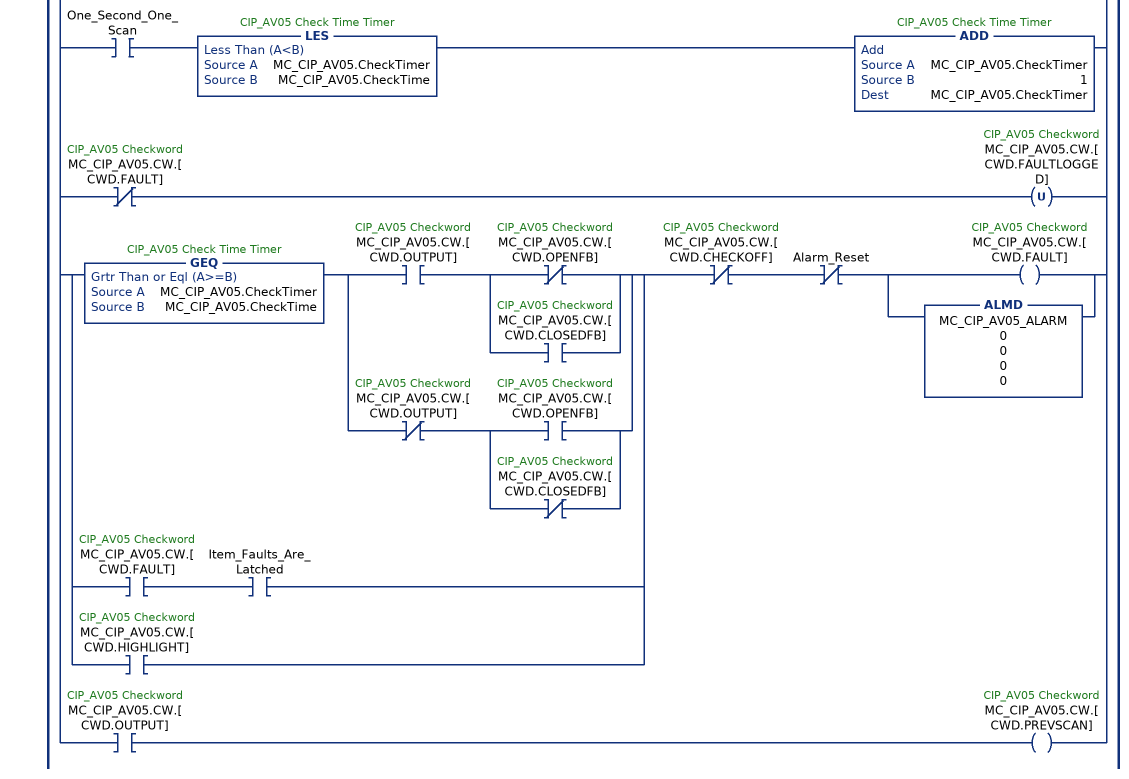
   62: [NEQ(MC_CIP_AV05.DriveBits,0) OTE(MC_CIP_AV05.CW.[CWD.AUTODRV]) ,[XIC(MC_CIP_AV05.CW.[CWD.AUTODRV]) XIO(MC_CIP_AV05.CW.[CWD.MANUAL]) ,XIC(MC_CIP_AV05.CW.[CWD.MANDRV]) XIC(MC_CIP_AV05.CW.[CWD.MANUAL]) ] OTE(MC_CIP_AV05.CW.[CWD.OUTPUT]) ,XIC(MC_CIP_AV05.CW.[CWD.OUTPUT]) OTE(MC_CIP_AV05_DR) ,XIC(S:FS) [OTU(MC_CIP_AV05.CW.[CWD.MANUAL]) ,LEQ(MC_CIP_AV05.CheckTime,0) MOV(Default_Check_Time,MC_CIP_AV05.CheckTime) ] ,[[XIC(MC_CIP_AV05_O) XIO(Item_Simulation_Flag) ,XIC(Item_Simulation_Flag) XIC(MC_CIP_AV05.CW.[CWD.OUTPUT]) XIO(MC_CIP_AV05.CW.[CWD.SIMFAIL]) ] OTE(MC_CIP_AV05.CW.[CWD.OPENFB]) ,[XIC(MC_CIP_AV05_C) XIO(Item_Simulation_Flag) ,XIC(Item_Simulation_Flag) XIO(MC_CIP_AV05.CW.[CWD.OUTPUT]) XIO(MC_CIP_AV05.CW.[CWD.SIMFAIL]) ] OTE(MC_CIP_AV05.CW.[CWD.CLOSEDFB]) ] ,[XIC(MC_CIP_AV05.CW.[CWD.OUTPUT]) XIO(MC_CIP_AV05.CW.[CWD.PREVSCAN]) ,XIO(MC_CIP_AV05.CW.[CWD.OUTPUT]) XIC(MC_CIP_AV05.CW.[CWD.PREVSCAN]) ] CLR(MC_CIP_AV05.CheckTimer) ,XIC(One_Second_One_Scan) LES(MC_CIP_AV05.CheckTimer,MC_CIP_AV05.CheckTime) ADD(MC_CIP_AV05.CheckTimer,1,MC_CIP_AV05.CheckTimer) ,XIO(MC_CIP_AV05.CW.[CWD.FAULT]) OTU(MC_CIP_AV05.CW.[CWD.FAULTLOGGED]) ,[GEQ(MC_CIP_AV05.CheckTimer,MC_CIP_AV05.CheckTime) [XIC(MC_CIP_AV05.CW.[CWD.OUTPUT]) [XIO(MC_CIP_AV05.CW.[CWD.OPENFB]) ,XIC(MC_CIP_AV05.CW.[CWD.CLOSEDFB]) ] ,XIO(MC_CIP_AV05.CW.[CWD.OUTPUT]) [XIC(MC_CIP_AV05.CW.[CWD.OPENFB]) ,XIO(MC_CIP_AV05.CW.[CWD.CLOSEDFB]) ] ] ,XIC(MC_CIP_AV05.CW.[CWD.FAULT]) XIC(Item_Faults_Are_Latched) ,XIC(MC_CIP_AV05.CW.[CWD.HIGHLIGHT]) ] XIO(MC_CIP_AV05.CW.[CWD.CHECKOFF]) XIO(Alarm_Reset) [OTE(MC_CIP_AV05.CW.[CWD.FAULT]) ,ALMD(MC_CIP_AV05_ALARM,0,0,0,0) ] ,XIC(MC_CIP_AV05.CW.[CWD.OUTPUT]) OTE(MC_CIP_AV05.CW.[CWD.PREVSCAN]) ];
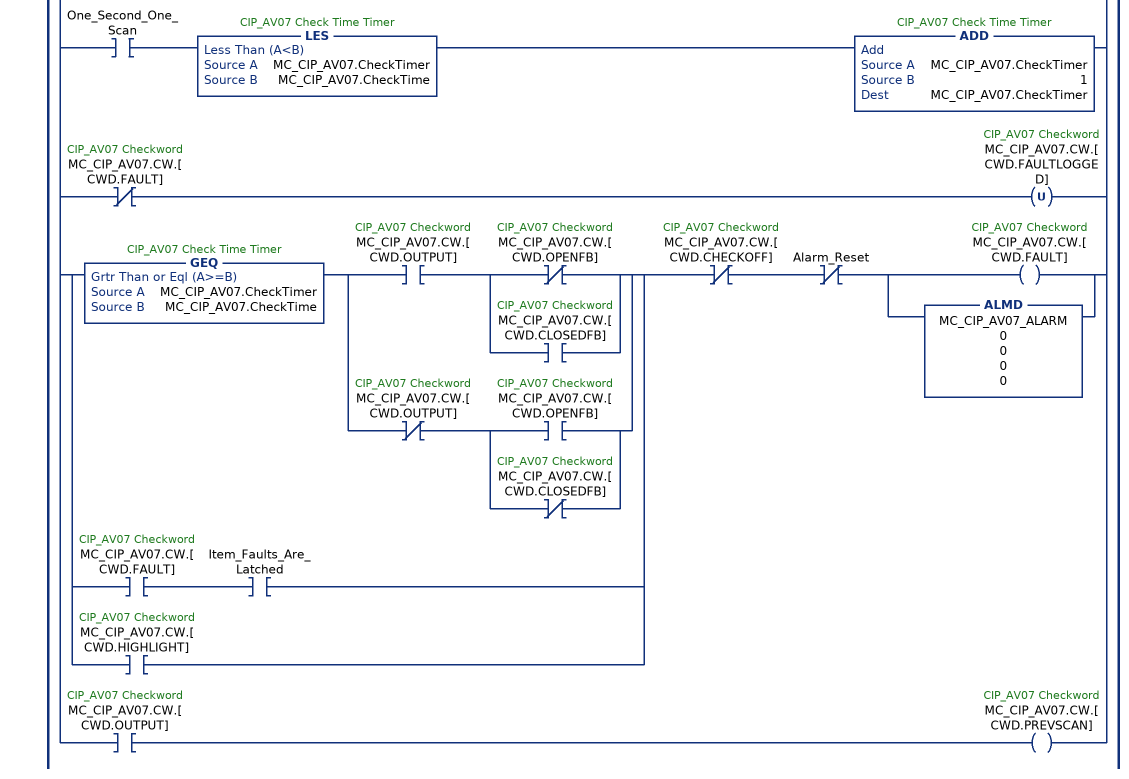
   63: [NEQ(MC_CIP_AV07.DriveBits,0) OTE(MC_CIP_AV07.CW.[CWD.AUTODRV]) ,[XIC(MC_CIP_AV07.CW.[CWD.AUTODRV]) XIO(MC_CIP_AV07.CW.[CWD.MANUAL]) ,XIC(MC_CIP_AV07.CW.[CWD.MANDRV]) XIC(MC_CIP_AV07.CW.[CWD.MANUAL]) ] OTE(MC_CIP_AV07.CW.[CWD.OUTPUT]) ,XIC(MC_CIP_AV07.CW.[CWD.OUTPUT]) OTE(MC_CIP_AV07_DR) ,XIC(S:FS) [OTU(MC_CIP_AV07.CW.[CWD.MANUAL]) ,LEQ(MC_CIP_AV07.CheckTime,0) MOV(Default_Check_Time,MC_CIP_AV07.CheckTime) ] ,[[XIC(MC_CIP_AV07_O) XIO(Item_Simulation_Flag) ,XIC(Item_Simulation_Flag) XIC(MC_CIP_AV07.CW.[CWD.OUTPUT]) XIO(MC_CIP_AV07.CW.[CWD.SIMFAIL]) ] OTE(MC_CIP_AV07.CW.[CWD.OPENFB]) ,[XIC(MC_CIP_AV07_C) XIO(Item_Simulation_Flag) ,XIC(Item_Simulation_Flag) XIO(MC_CIP_AV07.CW.[CWD.OUTPUT]) XIO(MC_CIP_AV07.CW.[CWD.SIMFAIL]) ] OTE(MC_CIP_AV07.CW.[CWD.CLOSEDFB]) ] ,[XIC(MC_CIP_AV07.CW.[CWD.OUTPUT]) XIO(MC_CIP_AV07.CW.[CWD.PREVSCAN]) ,XIO(MC_CIP_AV07.CW.[CWD.OUTPUT]) XIC(MC_CIP_AV07.CW.[CWD.PREVSCAN]) ] CLR(MC_CIP_AV07.CheckTimer) ,XIC(One_Second_One_Scan) LES(MC_CIP_AV07.CheckTimer,MC_CIP_AV07.CheckTime) ADD(MC_CIP_AV07.CheckTimer,1,MC_CIP_AV07.CheckTimer) ,XIO(MC_CIP_AV07.CW.[CWD.FAULT]) OTU(MC_CIP_AV07.CW.[CWD.FAULTLOGGED]) ,[GEQ(MC_CIP_AV07.CheckTimer,MC_CIP_AV07.CheckTime) [XIC(MC_CIP_AV07.CW.[CWD.OUTPUT]) [XIO(MC_CIP_AV07.CW.[CWD.OPENFB]) ,XIC(MC_CIP_AV07.CW.[CWD.CLOSEDFB]) ] ,XIO(MC_CIP_AV07.CW.[CWD.OUTPUT]) [XIC(MC_CIP_AV07.CW.[CWD.OPENFB]) ,XIO(MC_CIP_AV07.CW.[CWD.CLOSEDFB]) ] ] ,XIC(MC_CIP_AV07.CW.[CWD.FAULT]) XIC(Item_Faults_Are_Latched) ,XIC(MC_CIP_AV07.CW.[CWD.HIGHLIGHT]) ] XIO(MC_CIP_AV07.CW.[CWD.CHECKOFF]) XIO(Alarm_Reset) [OTE(MC_CIP_AV07.CW.[CWD.FAULT]) ,ALMD(MC_CIP_AV07_ALARM,0,0,0,0) ] ,XIC(MC_CIP_AV07.CW.[CWD.OUTPUT]) OTE(MC_CIP_AV07.CW.[CWD.PREVSCAN]) ];
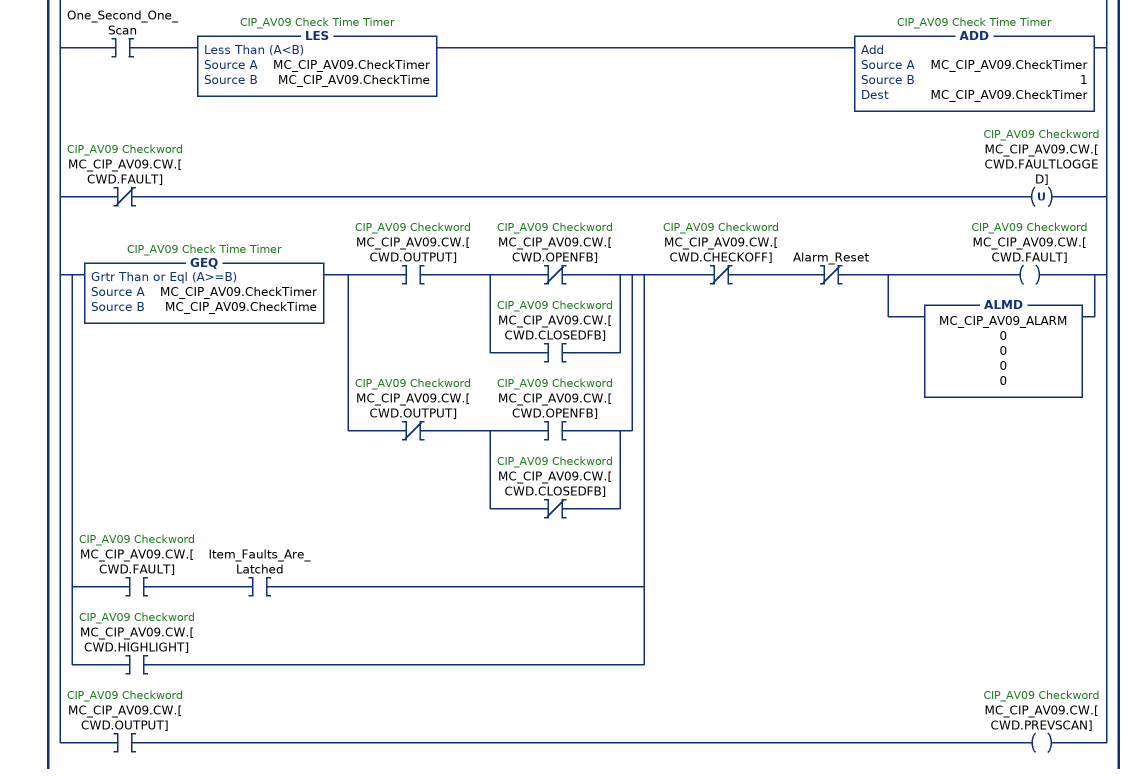
   64: [NEQ(MC_CIP_AV09.DriveBits,0) OTE(MC_CIP_AV09.CW.[CWD.AUTODRV]) ,[XIC(MC_CIP_AV09.CW.[CWD.AUTODRV]) XIO(MC_CIP_AV09.CW.[CWD.MANUAL]) ,XIC(MC_CIP_AV09.CW.[CWD.MANDRV]) XIC(MC_CIP_AV09.CW.[CWD.MANUAL]) ] OTE(MC_CIP_AV09.CW.[CWD.OUTPUT]) ,XIC(MC_CIP_AV09.CW.[CWD.OUTPUT]) OTE(MC_CIP_AV09_DR) ,XIC(S:FS) [OTU(MC_CIP_AV09.CW.[CWD.MANUAL]) ,LEQ(MC_CIP_AV09.CheckTime,0) MOV(Default_Check_Time,MC_CIP_AV09.CheckTime) ] ,[[XIC(MC_CIP_AV09_O) XIO(Item_Simulation_Flag) ,XIC(Item_Simulation_Flag) XIC(MC_CIP_AV09.CW.[CWD.OUTPUT]) XIO(MC_CIP_AV09.CW.[CWD.SIMFAIL]) ] OTE(MC_CIP_AV09.CW.[CWD.OPENFB]) ,[XIC(MC_CIP_AV09_C) XIO(Item_Simulation_Flag) ,XIC(Item_Simulation_Flag) XIO(MC_CIP_AV09.CW.[CWD.OUTPUT]) XIO(MC_CIP_AV09.CW.[CWD.SIMFAIL]) ] OTE(MC_CIP_AV09.CW.[CWD.CLOSEDFB]) ] ,[XIC(MC_CIP_AV09.CW.[CWD.OUTPUT]) XIO(MC_CIP_AV09.CW.[CWD.PREVSCAN]) ,XIO(MC_CIP_AV09.CW.[CWD.OUTPUT]) XIC(MC_CIP_AV09.CW.[CWD.PREVSCAN]) ] CLR(MC_CIP_AV09.CheckTimer) ,XIC(One_Second_One_Scan) LES(MC_CIP_AV09.CheckTimer,MC_CIP_AV09.CheckTime) ADD(MC_CIP_AV09.CheckTimer,1,MC_CIP_AV09.CheckTimer) ,XIO(MC_CIP_AV09.CW.[CWD.FAULT]) OTU(MC_CIP_AV09.CW.[CWD.FAULTLOGGED]) ,[GEQ(MC_CIP_AV09.CheckTimer,MC_CIP_AV09.CheckTime) [XIC(MC_CIP_AV09.CW.[CWD.OUTPUT]) [XIO(MC_CIP_AV09.CW.[CWD.OPENFB]) ,XIC(MC_CIP_AV09.CW.[CWD.CLOSEDFB]) ] ,XIO(MC_CIP_AV09.CW.[CWD.OUTPUT]) [XIC(MC_CIP_AV09.CW.[CWD.OPENFB]) ,XIO(MC_CIP_AV09.CW.[CWD.CLOSEDFB]) ] ] ,XIC(MC_CIP_AV09.CW.[CWD.FAULT]) XIC(Item_Faults_Are_Latched) ,XIC(MC_CIP_AV09.CW.[CWD.HIGHLIGHT]) ] XIO(MC_CIP_AV09.CW.[CWD.CHECKOFF]) XIO(Alarm_Reset) [OTE(MC_CIP_AV09.CW.[CWD.FAULT]) ,ALMD(MC_CIP_AV09_ALARM,0,0,0,0) ] ,XIC(MC_CIP_AV09.CW.[CWD.OUTPUT]) OTE(MC_CIP_AV09.CW.[CWD.PREVSCAN]) ];
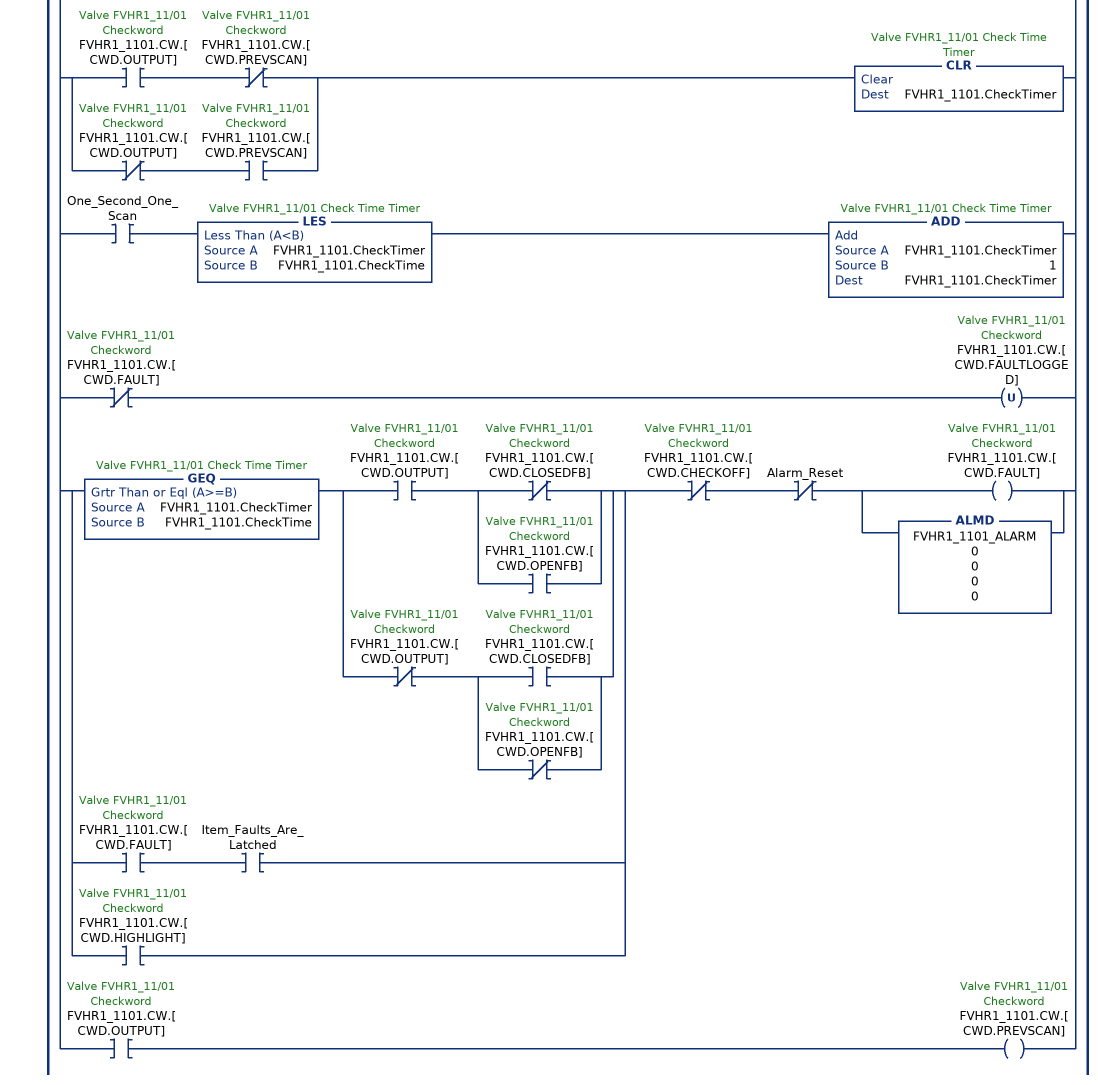
   65: [NEQ(FVHR1_1101.DriveBits,0) OTE(FVHR1_1101.CW.[CWD.AUTODRV]) ,[XIC(FVHR1_1101.CW.[CWD.AUTODRV]) XIO(FVHR1_1101.CW.[CWD.MANUAL]) ,XIC(FVHR1_1101.CW.[CWD.MANDRV]) XIC(FVHR1_1101.CW.[CWD.MANUAL]) ] OTE(FVHR1_1101.CW.[CWD.OUTPUT]) ,XIC(FVHR1_1101.CW.[CWD.OUTPUT]) OTE(FVHR1_1101_DR) ,XIC(S:FS) [OTU(FVHR1_1101.CW.[CWD.MANUAL]) ,LEQ(FVHR1_1101.CheckTime,0) MOV(Default_Check_Time,FVHR1_1101.CheckTime) ] ,[[XIC(FVHR1_1101_OP) XIO(Item_Simulation_Flag) ,XIC(Item_Simulation_Flag) XIC(FVHR1_1101.CW.[CWD.OUTPUT]) XIO(FVHR1_1101.CW.[CWD.SIMFAIL]) ] OTE(FVHR1_1101.CW.[CWD.OPENFB]) ,[XIC(FVHR1_1101_CL) XIO(Item_Simulation_Flag) ,XIC(Item_Simulation_Flag) XIO(FVHR1_1101.CW.[CWD.OUTPUT]) XIO(FVHR1_1101.CW.[CWD.SIMFAIL]) ] OTE(FVHR1_1101.CW.[CWD.CLOSEDFB]) ] ,[XIC(FVHR1_1101.CW.[CWD.OUTPUT]) XIO(FVHR1_1101.CW.[CWD.PREVSCAN]) ,XIO(FVHR1_1101.CW.[CWD.OUTPUT]) XIC(FVHR1_1101.CW.[CWD.PREVSCAN]) ] CLR(FVHR1_1101.CheckTimer) ,XIC(One_Second_One_Scan) LES(FVHR1_1101.CheckTimer,FVHR1_1101.CheckTime) ADD(FVHR1_1101.CheckTimer,1,FVHR1_1101.CheckTimer) ,XIO(FVHR1_1101.CW.[CWD.FAULT]) OTU(FVHR1_1101.CW.[CWD.FAULTLOGGED]) ,[GEQ(FVHR1_1101.CheckTimer,FVHR1_1101.CheckTime) [XIC(FVHR1_1101.CW.[CWD.OUTPUT]) [XIO(FVHR1_1101.CW.[CWD.CLOSEDFB]) ,XIC(FVHR1_1101.CW.[CWD.OPENFB]) ] ,XIO(FVHR1_1101.CW.[CWD.OUTPUT]) [XIC(FVHR1_1101.CW.[CWD.CLOSEDFB]) ,XIO(FVHR1_1101.CW.[CWD.OPENFB]) ] ] ,XIC(FVHR1_1101.CW.[CWD.FAULT]) XIC(Item_Faults_Are_Latched) ,XIC(FVHR1_1101.CW.[CWD.HIGHLIGHT]) ] XIO(FVHR1_1101.CW.[CWD.CHECKOFF]) XIO(Alarm_Reset) [OTE(FVHR1_1101.CW.[CWD.FAULT]) ,ALMD(FVHR1_1101_ALARM,0,0,0,0) ] ,XIC(FVHR1_1101.CW.[CWD.OUTPUT]) OTE(FVHR1_1101.CW.[CWD.PREVSCAN]) ];
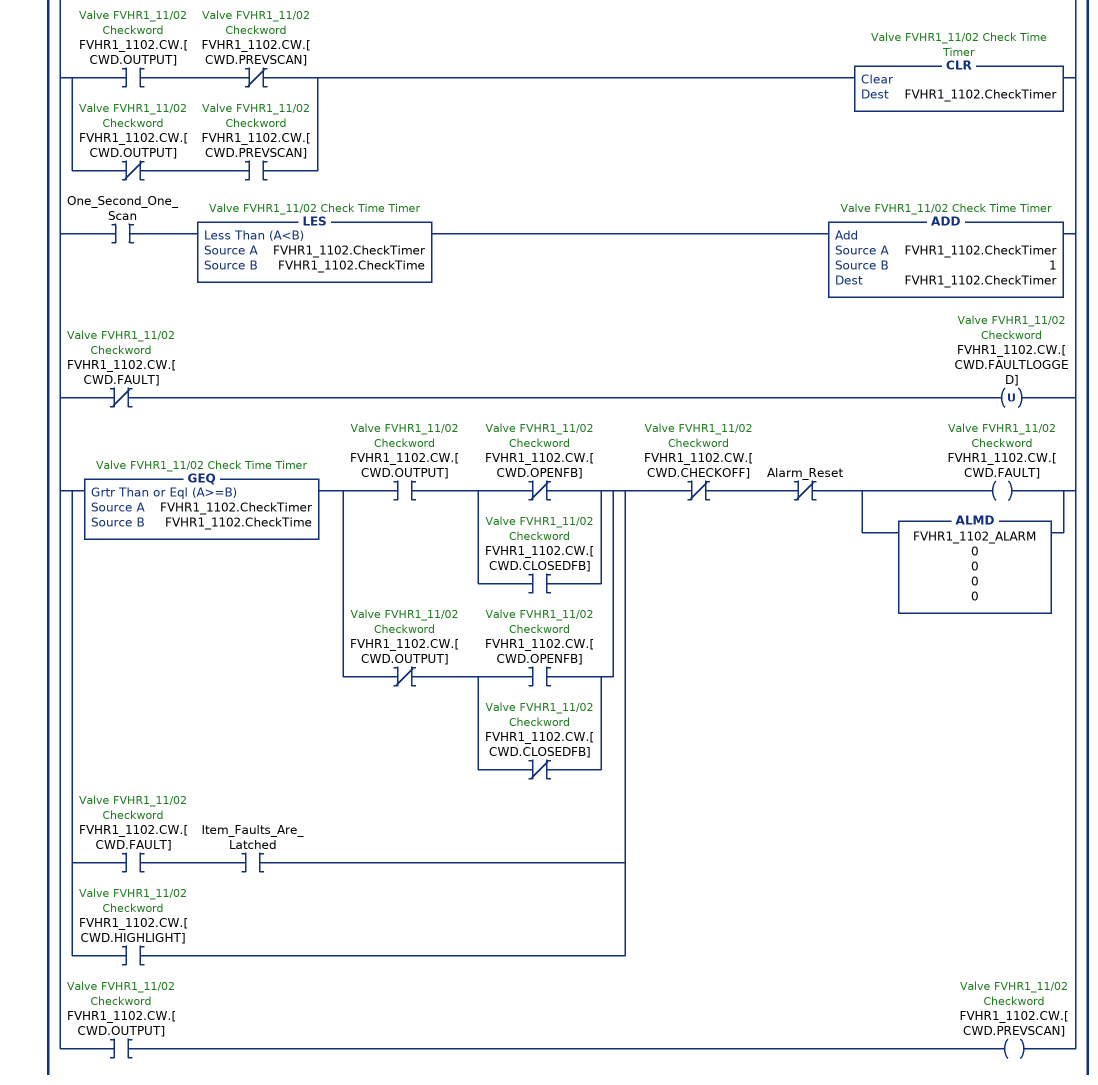
   66: [NEQ(FVHR1_1102.DriveBits,0) OTE(FVHR1_1102.CW.[CWD.AUTODRV]) ,[XIC(FVHR1_1102.CW.[CWD.AUTODRV]) XIO(FVHR1_1102.CW.[CWD.MANUAL]) ,XIC(FVHR1_1102.CW.[CWD.MANDRV]) XIC(FVHR1_1102.CW.[CWD.MANUAL]) ] OTE(FVHR1_1102.CW.[CWD.OUTPUT]) ,XIC(FVHR1_1102.CW.[CWD.OUTPUT]) OTE(FVHR1_1102_DR) ,XIC(S:FS) [OTU(FVHR1_1102.CW.[CWD.MANUAL]) ,LEQ(FVHR1_1102.CheckTime,0) MOV(Default_Check_Time,FVHR1_1102.CheckTime) ] ,[[XIC(FVHR1_1102_OP) XIO(Item_Simulation_Flag) ,XIC(Item_Simulation_Flag) XIC(FVHR1_1102.CW.[CWD.OUTPUT]) XIO(FVHR1_1102.CW.[CWD.SIMFAIL]) ] OTE(FVHR1_1102.CW.[CWD.OPENFB]) ,[XIC(FVHR1_1102_CL) XIO(Item_Simulation_Flag) ,XIC(Item_Simulation_Flag) XIO(FVHR1_1102.CW.[CWD.OUTPUT]) XIO(FVHR1_1102.CW.[CWD.SIMFAIL]) ] OTE(FVHR1_1102.CW.[CWD.CLOSEDFB]) ] ,[XIC(FVHR1_1102.CW.[CWD.OUTPUT]) XIO(FVHR1_1102.CW.[CWD.PREVSCAN]) ,XIO(FVHR1_1102.CW.[CWD.OUTPUT]) XIC(FVHR1_1102.CW.[CWD.PREVSCAN]) ] CLR(FVHR1_1102.CheckTimer) ,XIC(One_Second_One_Scan) LES(FVHR1_1102.CheckTimer,FVHR1_1102.CheckTime) ADD(FVHR1_1102.CheckTimer,1,FVHR1_1102.CheckTimer) ,XIO(FVHR1_1102.CW.[CWD.FAULT]) OTU(FVHR1_1102.CW.[CWD.FAULTLOGGED]) ,[GEQ(FVHR1_1102.CheckTimer,FVHR1_1102.CheckTime) [XIC(FVHR1_1102.CW.[CWD.OUTPUT]) [XIO(FVHR1_1102.CW.[CWD.OPENFB]) ,XIC(FVHR1_1102.CW.[CWD.CLOSEDFB]) ] ,XIO(FVHR1_1102.CW.[CWD.OUTPUT]) [XIC(FVHR1_1102.CW.[CWD.OPENFB]) ,XIO(FVHR1_1102.CW.[CWD.CLOSEDFB]) ] ] ,XIC(FVHR1_1102.CW.[CWD.FAULT]) XIC(Item_Faults_Are_Latched) ,XIC(FVHR1_1102.CW.[CWD.HIGHLIGHT]) ] XIO(FVHR1_1102.CW.[CWD.CHECKOFF]) XIO(Alarm_Reset) [OTE(FVHR1_1102.CW.[CWD.FAULT]) ,ALMD(FVHR1_1102_ALARM,0,0,0,0) ] ,XIC(FVHR1_1102.CW.[CWD.OUTPUT]) OTE(FVHR1_1102.CW.[CWD.PREVSCAN]) ];
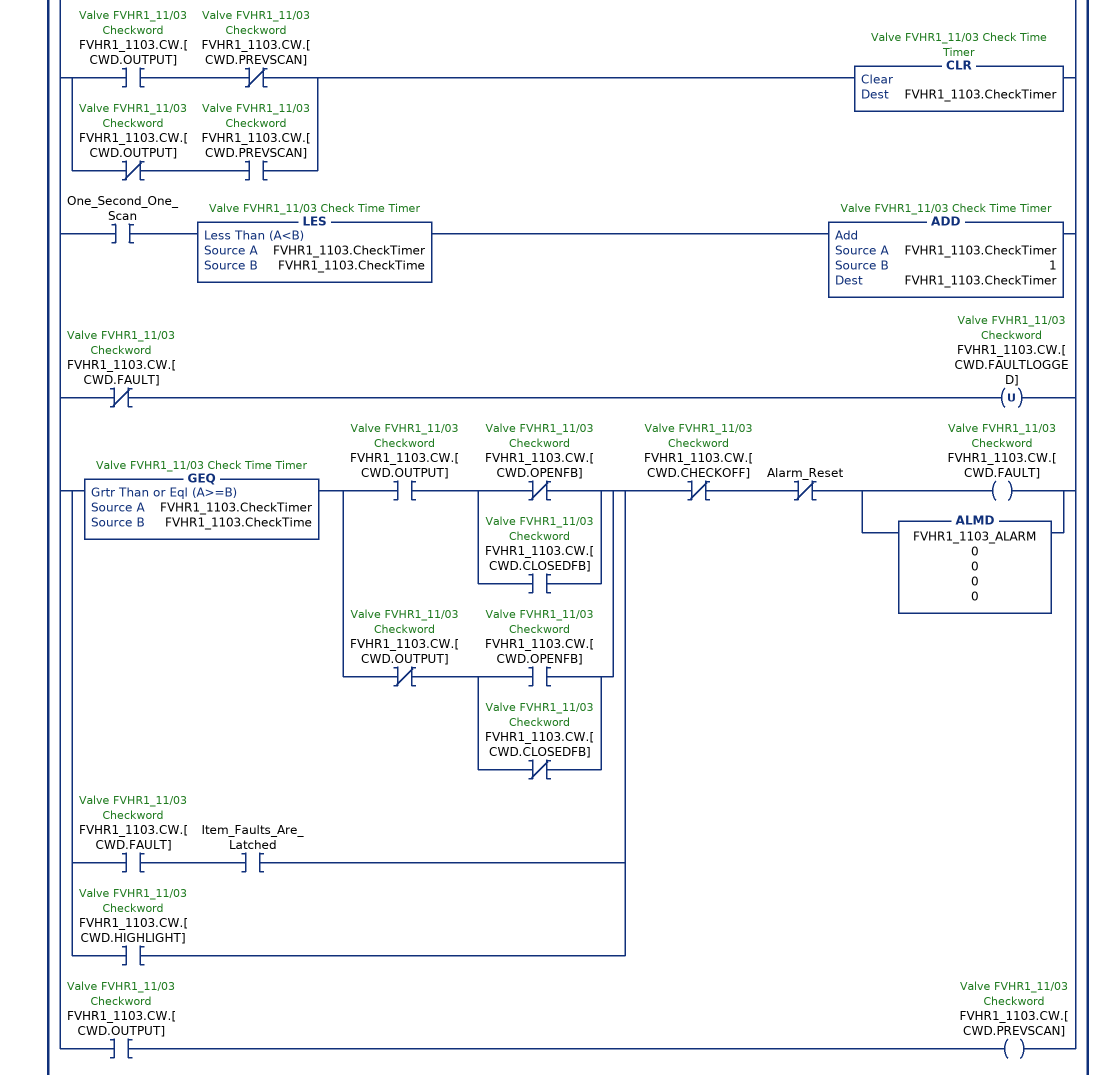
   67: [NEQ(FVHR1_1103.DriveBits,0) OTE(FVHR1_1103.CW.[CWD.AUTODRV]) ,[XIC(FVHR1_1103.CW.[CWD.AUTODRV]) XIO(FVHR1_1103.CW.[CWD.MANUAL]) ,XIC(FVHR1_1103.CW.[CWD.MANDRV]) XIC(FVHR1_1103.CW.[CWD.MANUAL]) ] OTE(FVHR1_1103.CW.[CWD.OUTPUT]) ,XIC(FVHR1_1103.CW.[CWD.OUTPUT]) OTE(FVHR1_1103_DR) ,XIC(S:FS) [OTU(FVHR1_1103.CW.[CWD.MANUAL]) ,LEQ(FVHR1_1103.CheckTime,0) MOV(Default_Check_Time,FVHR1_1103.CheckTime) ] ,[[XIC(FVHR1_1103_OP) XIO(Item_Simulation_Flag) ,XIC(Item_Simulation_Flag) XIC(FVHR1_1103.CW.[CWD.OUTPUT]) XIO(FVHR1_1103.CW.[CWD.SIMFAIL]) ] OTE(FVHR1_1103.CW.[CWD.OPENFB]) ,[XIC(FVHR1_1103_CL) XIO(Item_Simulation_Flag) ,XIC(Item_Simulation_Flag) XIO(FVHR1_1103.CW.[CWD.OUTPUT]) XIO(FVHR1_1103.CW.[CWD.SIMFAIL]) ] OTE(FVHR1_1103.CW.[CWD.CLOSEDFB]) ] ,[XIC(FVHR1_1103.CW.[CWD.OUTPUT]) XIO(FVHR1_1103.CW.[CWD.PREVSCAN]) ,XIO(FVHR1_1103.CW.[CWD.OUTPUT]) XIC(FVHR1_1103.CW.[CWD.PREVSCAN]) ] CLR(FVHR1_1103.CheckTimer) ,XIC(One_Second_One_Scan) LES(FVHR1_1103.CheckTimer,FVHR1_1103.CheckTime) ADD(FVHR1_1103.CheckTimer,1,FVHR1_1103.CheckTimer) ,XIO(FVHR1_1103.CW.[CWD.FAULT]) OTU(FVHR1_1103.CW.[CWD.FAULTLOGGED]) ,[GEQ(FVHR1_1103.CheckTimer,FVHR1_1103.CheckTime) [XIC(FVHR1_1103.CW.[CWD.OUTPUT]) [XIO(FVHR1_1103.CW.[CWD.OPENFB]) ,XIC(FVHR1_1103.CW.[CWD.CLOSEDFB]) ] ,XIO(FVHR1_1103.CW.[CWD.OUTPUT]) [XIC(FVHR1_1103.CW.[CWD.OPENFB]) ,XIO(FVHR1_1103.CW.[CWD.CLOSEDFB]) ] ] ,XIC(FVHR1_1103.CW.[CWD.FAULT]) XIC(Item_Faults_Are_Latched) ,XIC(FVHR1_1103.CW.[CWD.HIGHLIGHT]) ] XIO(FVHR1_1103.CW.[CWD.CHECKOFF]) XIO(Alarm_Reset) [OTE(FVHR1_1103.CW.[CWD.FAULT]) ,ALMD(FVHR1_1103_ALARM,0,0,0,0) ] ,XIC(FVHR1_1103.CW.[CWD.OUTPUT]) OTE(FVHR1_1103.CW.[CWD.PREVSCAN]) ];
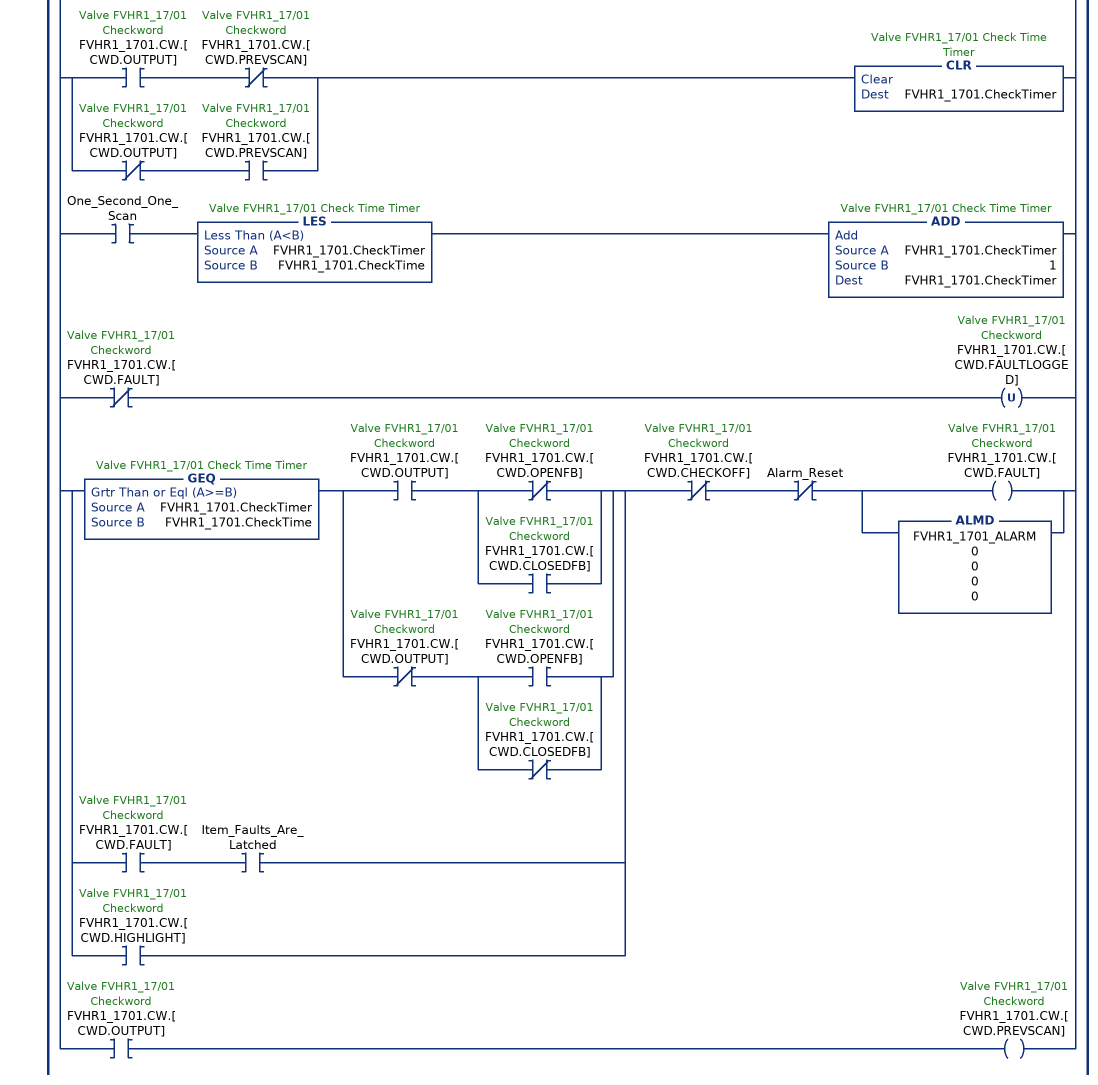
   68: [NEQ(FVHR1_1701.DriveBits,0) OTE(FVHR1_1701.CW.[CWD.AUTODRV]) ,[XIC(FVHR1_1701.CW.[CWD.AUTODRV]) XIO(FVHR1_1701.CW.[CWD.MANUAL]) ,XIC(FVHR1_1701.CW.[CWD.MANDRV]) XIC(FVHR1_1701.CW.[CWD.MANUAL]) ] OTE(FVHR1_1701.CW.[CWD.OUTPUT]) ,XIC(FVHR1_1701.CW.[CWD.OUTPUT]) OTE(FVHR1_1701_DR) ,XIC(S:FS) [OTU(FVHR1_1701.CW.[CWD.MANUAL]) ,LEQ(FVHR1_1701.CheckTime,0) MOV(Default_Check_Time,FVHR1_1701.CheckTime) ] ,[[XIC(FVHR1_1701_OP) XIO(Item_Simulation_Flag) ,XIC(Item_Simulation_Flag) XIC(FVHR1_1701.CW.[CWD.OUTPUT]) XIO(FVHR1_1701.CW.[CWD.SIMFAIL]) ] OTE(FVHR1_1701.CW.[CWD.OPENFB]) ,[XIC(FVHR1_1701_CL) XIO(Item_Simulation_Flag) ,XIC(Item_Simulation_Flag) XIO(FVHR1_1701.CW.[CWD.OUTPUT]) XIO(FVHR1_1701.CW.[CWD.SIMFAIL]) ] OTE(FVHR1_1701.CW.[CWD.CLOSEDFB]) ] ,[XIC(FVHR1_1701.CW.[CWD.OUTPUT]) XIO(FVHR1_1701.CW.[CWD.PREVSCAN]) ,XIO(FVHR1_1701.CW.[CWD.OUTPUT]) XIC(FVHR1_1701.CW.[CWD.PREVSCAN]) ] CLR(FVHR1_1701.CheckTimer) ,XIC(One_Second_One_Scan) LES(FVHR1_1701.CheckTimer,FVHR1_1701.CheckTime) ADD(FVHR1_1701.CheckTimer,1,FVHR1_1701.CheckTimer) ,XIO(FVHR1_1701.CW.[CWD.FAULT]) OTU(FVHR1_1701.CW.[CWD.FAULTLOGGED]) ,[GEQ(FVHR1_1701.CheckTimer,FVHR1_1701.CheckTime) [XIC(FVHR1_1701.CW.[CWD.OUTPUT]) [XIO(FVHR1_1701.CW.[CWD.OPENFB]) ,XIC(FVHR1_1701.CW.[CWD.CLOSEDFB]) ] ,XIO(FVHR1_1701.CW.[CWD.OUTPUT]) [XIC(FVHR1_1701.CW.[CWD.OPENFB]) ,XIO(FVHR1_1701.CW.[CWD.CLOSEDFB]) ] ] ,XIC(FVHR1_1701.CW.[CWD.FAULT]) XIC(Item_Faults_Are_Latched) ,XIC(FVHR1_1701.CW.[CWD.HIGHLIGHT]) ] XIO(FVHR1_1701.CW.[CWD.CHECKOFF]) XIO(Alarm_Reset) [OTE(FVHR1_1701.CW.[CWD.FAULT]) ,ALMD(FVHR1_1701_ALARM,0,0,0,0) ] ,XIC(FVHR1_1701.CW.[CWD.OUTPUT]) OTE(FVHR1_1701.CW.[CWD.PREVSCAN]) ];
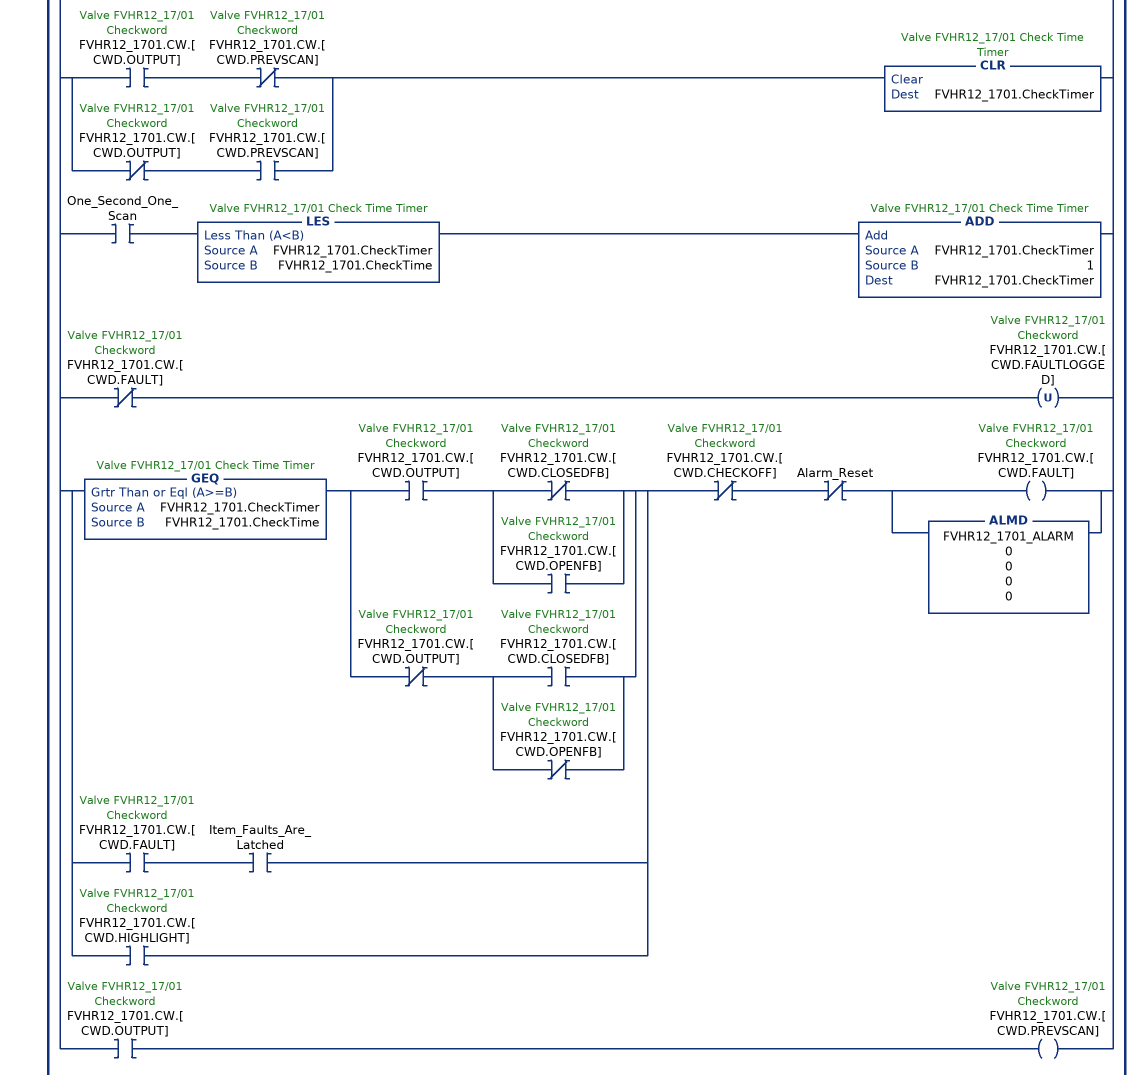
   69: [NEQ(FVHR12_1701.DriveBits,0) OTE(FVHR12_1701.CW.[CWD.AUTODRV]) ,[XIC(FVHR12_1701.CW.[CWD.AUTODRV]) XIO(FVHR12_1701.CW.[CWD.MANUAL]) ,XIC(FVHR12_1701.CW.[CWD.MANDRV]) XIC(FVHR12_1701.CW.[CWD.MANUAL]) ] OTE(FVHR12_1701.CW.[CWD.OUTPUT]) ,XIC(FVHR12_1701.CW.[CWD.OUTPUT]) OTE(FVHR12_1701_DR) ,XIC(S:FS) [OTU(FVHR12_1701.CW.[CWD.MANUAL]) ,LEQ(FVHR12_1701.CheckTime,0) MOV(Default_Check_Time,FVHR12_1701.CheckTime) ] ,[[XIC(FVHR12_1701_OP) XIO(Item_Simulation_Flag) ,XIC(Item_Simulation_Flag) XIC(FVHR12_1701.CW.[CWD.OUTPUT]) XIO(FVHR12_1701.CW.[CWD.SIMFAIL]) ] OTE(FVHR12_1701.CW.[CWD.OPENFB]) ,[XIC(FVHR12_1701_CL) XIO(Item_Simulation_Flag) ,XIC(Item_Simulation_Flag) XIO(FVHR12_1701.CW.[CWD.OUTPUT]) XIO(FVHR12_1701.CW.[CWD.SIMFAIL]) ] OTE(FVHR12_1701.CW.[CWD.CLOSEDFB]) ] ,[XIC(FVHR12_1701.CW.[CWD.OUTPUT]) XIO(FVHR12_1701.CW.[CWD.PREVSCAN]) ,XIO(FVHR12_1701.CW.[CWD.OUTPUT]) XIC(FVHR12_1701.CW.[CWD.PREVSCAN]) ] CLR(FVHR12_1701.CheckTimer) ,XIC(One_Second_One_Scan) LES(FVHR12_1701.CheckTimer,FVHR12_1701.CheckTime) ADD(FVHR12_1701.CheckTimer,1,FVHR12_1701.CheckTimer) ,XIO(FVHR12_1701.CW.[CWD.FAULT]) OTU(FVHR12_1701.CW.[CWD.FAULTLOGGED]) ,[GEQ(FVHR12_1701.CheckTimer,FVHR12_1701.CheckTime) [XIC(FVHR12_1701.CW.[CWD.OUTPUT]) [XIO(FVHR12_1701.CW.[CWD.CLOSEDFB]) ,XIC(FVHR12_1701.CW.[CWD.OPENFB]) ] ,XIO(FVHR12_1701.CW.[CWD.OUTPUT]) [XIC(FVHR12_1701.CW.[CWD.CLOSEDFB]) ,XIO(FVHR12_1701.CW.[CWD.OPENFB]) ] ] ,XIC(FVHR12_1701.CW.[CWD.FAULT]) XIC(Item_Faults_Are_Latched) ,XIC(FVHR12_1701.CW.[CWD.HIGHLIGHT]) ] XIO(FVHR12_1701.CW.[CWD.CHECKOFF]) XIO(Alarm_Reset) [OTE(FVHR12_1701.CW.[CWD.FAULT]) ,ALMD(FVHR12_1701_ALARM,0,0,0,0) ] ,XIC(FVHR12_1701.CW.[CWD.OUTPUT]) OTE(FVHR12_1701.CW.[CWD.PREVSCAN]) ];
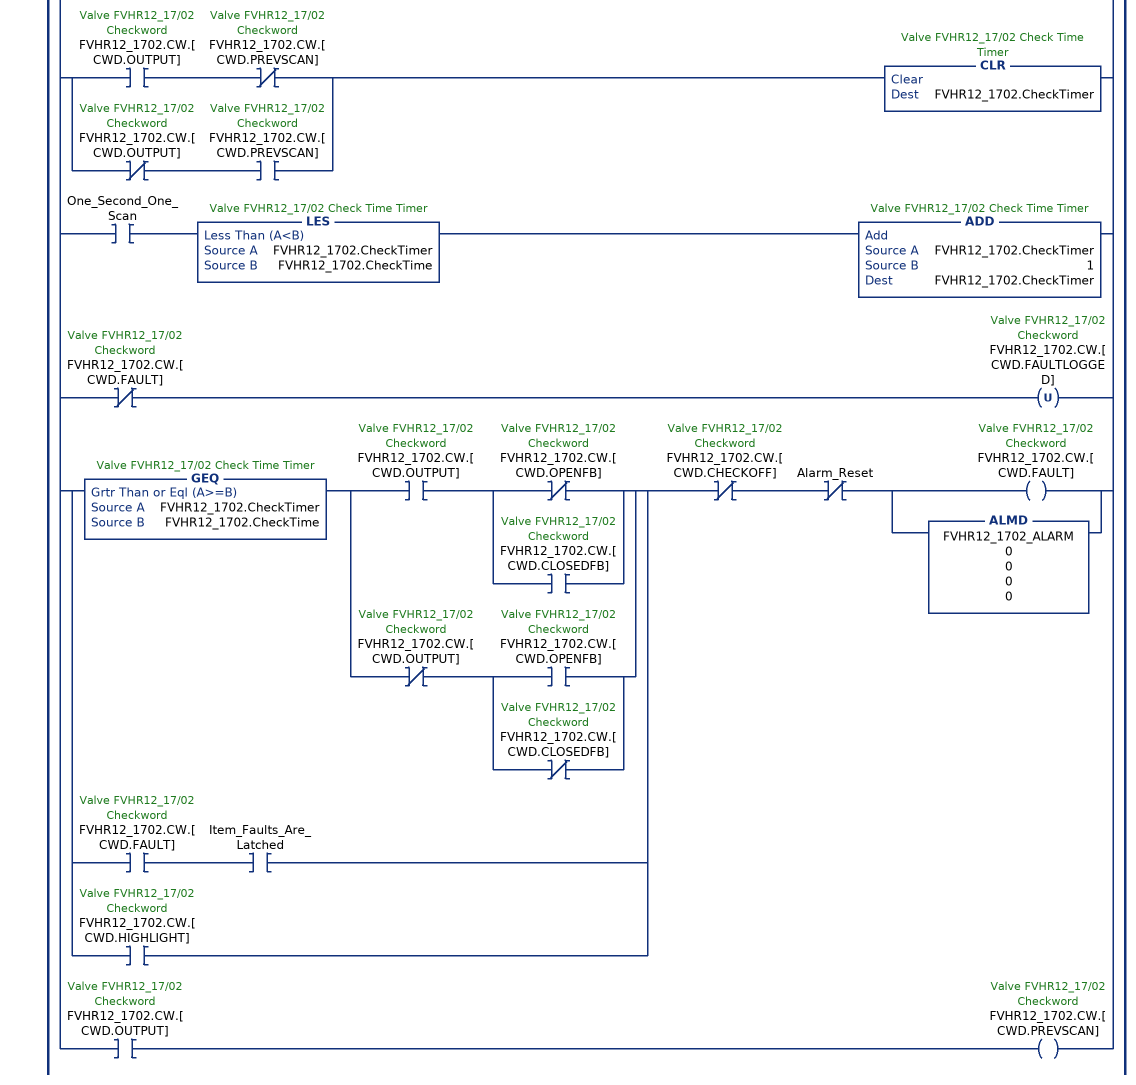
   70: [NEQ(FVHR12_1702.DriveBits,0) OTE(FVHR12_1702.CW.[CWD.AUTODRV]) ,[XIC(FVHR12_1702.CW.[CWD.AUTODRV]) XIO(FVHR12_1702.CW.[CWD.MANUAL]) ,XIC(FVHR12_1702.CW.[CWD.MANDRV]) XIC(FVHR12_1702.CW.[CWD.MANUAL]) ] OTE(FVHR12_1702.CW.[CWD.OUTPUT]) ,XIC(FVHR12_1702.CW.[CWD.OUTPUT]) OTE(FVHR12_1702_DR) ,XIC(S:FS) [OTU(FVHR12_1702.CW.[CWD.MANUAL]) ,LEQ(FVHR12_1702.CheckTime,0) MOV(Default_Check_Time,FVHR12_1702.CheckTime) ] ,[[XIC(FVHR12_1702_OP) XIO(Item_Simulation_Flag) ,XIC(Item_Simulation_Flag) XIC(FVHR12_1702.CW.[CWD.OUTPUT]) XIO(FVHR12_1702.CW.[CWD.SIMFAIL]) ] OTE(FVHR12_1702.CW.[CWD.OPENFB]) ,[XIC(FVHR12_1702_CL) XIO(Item_Simulation_Flag) ,XIC(Item_Simulation_Flag) XIO(FVHR12_1702.CW.[CWD.OUTPUT]) XIO(FVHR12_1702.CW.[CWD.SIMFAIL]) ] OTE(FVHR12_1702.CW.[CWD.CLOSEDFB]) ] ,[XIC(FVHR12_1702.CW.[CWD.OUTPUT]) XIO(FVHR12_1702.CW.[CWD.PREVSCAN]) ,XIO(FVHR12_1702.CW.[CWD.OUTPUT]) XIC(FVHR12_1702.CW.[CWD.PREVSCAN]) ] CLR(FVHR12_1702.CheckTimer) ,XIC(One_Second_One_Scan) LES(FVHR12_1702.CheckTimer,FVHR12_1702.CheckTime) ADD(FVHR12_1702.CheckTimer,1,FVHR12_1702.CheckTimer) ,XIO(FVHR12_1702.CW.[CWD.FAULT]) OTU(FVHR12_1702.CW.[CWD.FAULTLOGGED]) ,[GEQ(FVHR12_1702.CheckTimer,FVHR12_1702.CheckTime) [XIC(FVHR12_1702.CW.[CWD.OUTPUT]) [XIO(FVHR12_1702.CW.[CWD.OPENFB]) ,XIC(FVHR12_1702.CW.[CWD.CLOSEDFB]) ] ,XIO(FVHR12_1702.CW.[CWD.OUTPUT]) [XIC(FVHR12_1702.CW.[CWD.OPENFB]) ,XIO(FVHR12_1702.CW.[CWD.CLOSEDFB]) ] ] ,XIC(FVHR12_1702.CW.[CWD.FAULT]) XIC(Item_Faults_Are_Latched) ,XIC(FVHR12_1702.CW.[CWD.HIGHLIGHT]) ] XIO(FVHR12_1702.CW.[CWD.CHECKOFF]) XIO(Alarm_Reset) [OTE(FVHR12_1702.CW.[CWD.FAULT]) ,ALMD(FVHR12_1702_ALARM,0,0,0,0) ] ,XIC(FVHR12_1702.CW.[CWD.OUTPUT]) OTE(FVHR12_1702.CW.[CWD.PREVSCAN]) ];